   TextField "Text field_116" at 102,429 size 382x38; Text 'Tank 1P GTT Isolation Valve Feedback - Opened CV422'
   TextField "Text field_117" at 102,465 size 374x38; Text 'Tank 1P GTT Isolation Valve Feedback - Closed CV422'
   TextField "Text field_118" at 102,501 size 371x38; Text 'Tank 1P Tank Vent Valve 1 Feedback - Opened CV441-1PA'
   TextField "Text field_119" at 102,537 size 363x38; Text 'Tank 1P Tank Vent Valve 1 Feedback - Closed CV441-1PA'
   TextField "Text field_120" at 102,573 size 371x38; Text 'Tank 1P Tank Vent Valve 2 Feedback - Opened CV441-1PB'
   TextField "Text field_121" at 102,609 size 363x38; Text 'Tank 1P Tank Vent Valve 2 Feedback - Closed CV441-1PB'
   TextField "Text field_122" at 102,690 size 100x21; Text 'Spare Input'
   TextField "Text field_123" at 636,113 size 382x38; Text 'Tank 1S GTT Isolation Valve Feedback - Opened CV421'
   TextField "Text field_124" at 636,148 size 374x38; Text 'Tank 1S GTT Isolation Valve Feedback - Closed CV421'
   TextField "Text field_125" at 636,184 size 371x38; Text 'Tank 1S Tank Vent Valve 1 Feedback - Opened CV440-1SA'
   TextField "Text field_126" at 636,219 size 363x38; Text 'Tank 1S Tank Vent Valve 1 Feedback - Closed CV440-1SA'
   TextField "Text field_127" at 636,255 size 371x38; Text 'Tank 1S Tank Vent Valve 2 Feedback - Opened CV440-1SB'
   TextField "Text field_128" at 636,291 size 363x38; Text 'Tank 1S Tank Vent Valve 2 Feedback - Closed CV440-1SB'
   TextField "Text field_129" at 636,328 size 100x21; Text 'Spare Input'
   TextField "Text field_130" at 636,366 size 100x21; Text 'Spare Input'
   TextField "Text field_131" at 635,431 size 260x38; Text 'FPT BWT Level High High Switch LS425-FPT'
   TextField "Text field_132" at 635,467 size 270x38; Text 'RIO1 Tanks Pressure Switch Hi Hi PS436-FPT/1P/1S'
   TextField "Text field_133" at 635,503 size 294x38; Text 'Tank 1P BWT Level High High Switch LS425-1P'
   TextField "Text field_134" at 635,611 size 100x21; Text 'Spare Input'
   TextField "Text field_135" at 635,648 size 100x21; Text 'Spare Input'
   TextField "Text field_136" at 635,688 size 100x21; Text 'Spare Input'
   TextField "Text field_137" at 635,539 size 294x38; Text 'Tank 1S BWT Level High High Switch LS425-1S'
   TextField "Text field_138" at 635,576 size 100x21; Text 'Spare Input'
   TextField "Text field_115" at 102,654 size 100x21; Text 'Spare Input'
   AlarmView "Alarm view_1" at 0,777 size 1280x23
   Group "Group" at 455,41 size 373x50
   Button "HmiScreenItemData_8" at 469,45 size 355x40; TextOn 'Back'; TextOff 'Text'
      on Click: "TitleUpdater"()
   TextField "Screen title" at 455,41 size 373x50; Text 'Screen title'

screen "IGG Digital Outputs" 1280x800, template "Template"
   on GenerateScreen: "TitleUpdater"()
   Button "HmiScreenItemData_1" at 1,1 size 150x43; TextOn 'Back'; TextOff 'Commissioning'
      on Release: ActivateScreen("Commissioning Main Page", 0)
   AlarmView "Alarm view_1" at 0,777 size 1280x23
   TextField "Text field_1" at 395,239 size 55x22; Text 'Q0.0'
   TextField "Text field_2" at 395,290 size 55x22; Text 'Q0.1'
   TextField "Text field_3" at 395,342 size 55x22; Text 'Q0.2'
   TextField "Text field_4" at 395,394 size 55x22; Text 'Q0.3'
   TextField "Text field_5" at 395,446 size 55x22; Text 'Q0.4'
   TextField "Text field_6" at 395,498 size 55x22; Text 'Q0.5'
   TextField "Text field_7" at 395,550 size 55x22; Text 'Q0.6'
   TextField "Text field_8" at 395,602 size 55x22; Text 'Q0.7'
   Circle "Circle_1" at 455,239 size 20x20
      Appearance <- "14_DQ_Data_E500A_CNTRL"
   Circle "Circle_2" at 455,290 size 20x20
      Appearance <- "14_DQ_Data_E500B_CNTRL"
   Circle "Circle_3" at 455,342 size 20x20
      Appearance <- "14_DQ_Data_E139_CNTRL"
   Circle "Circle_4" at 455,394 size 20x20
      Appearance <- "14_DQ_Data_CV311_312_CNTRL"
   Circle "Circle_5" at 455,446 size 20x20
      Appearance <- "14_DQ_Data_CV321_322_CNTRL"
   Circle "Circle_6" at 455,498 size 20x20
      Appearance <- "14_DQ_Data_CV401_CNTRL"
   Circle "Circle_7" at 455,550 size 20x20
      Appearance <- "14_DQ_Data_CV431_432_CNTRL"
   Circle "Circle_8" at 455,602 size 20x20
      Appearance <- "14_DQ_Data_R2_SPR_DQ_0_7"
   TextField "Text field_9" at 412,206 size 49x26; Text 'Q0'
   TextField "Text field_10" at 698,239 size 55x22; Text 'Q1.0'
   TextField "Text field_11" at 698,290 size 55x22; Text 'Q1.1'
   TextField "Text field_12" at 698,342 size 55x22; Text 'Q1.2'
   TextField "Text field_13" at 698,394 size 55x22; Text 'Q1.3'
   TextField "Text field_14" at 698,446 size 55x22; Text 'Q1.4'
   TextField "Text field_15" at 698,498 size 55x22; Text 'Q1.5'
   TextField "Text field_16" at 698,550 size 55x22; Text 'Q1.6'
   TextField "Text field_17" at 698,602 size 55x22; Text 'Q1.7'
   Circle "Circle_9" at 758,239 size 20x20
      Appearance <- "14_DQ_Data_R2_SPR_DQ_1_0"
   Circle "Circle_10" at 758,290 size 20x20
      Appearance <- "14_DQ_Data_24K2"
   Circle "Circle_11" at 758,342 size 20x20
      Appearance <- "14_DQ_Data_24K3"
   Circle "Circle_12" at 758,394 size 20x20
      Appearance <- "14_DQ_Data_24K4"
   Circle "Circle_13" at 758,446 size 20x20
      Appearance <- "14_DQ_Data_24PF1"
   Circle "Circle_14" at 758,498 size 20x20
      Appearance <- "14_DQ_Data_24PF2"
   Circle "Circle_15" at 758,550 size 20x20
      Appearance <- "14_DQ_Data_24PF3"
   Circle "Circle_16" at 758,602 size 20x20
      Appearance <- "14_DQ_Data_24PF4"
   TextField "Text field_18" at 715,206 size 49x26; Text 'Q1'
   TextField "Text field_37" at 328,167 size 254x26; Text 'IGG System PLC (Rack 1)'
   Button "Button_9" at 330,493 size 60x35; TextOff 'Override'
      on Press: InvertBit("80_From_HMI_MAN_DQ_0_5")
      Visibility <- "82_To_HMI_CRNT_MODE_IGG"
   Button "Button_10" at 330,441 size 60x35; TextOff 'Override'
      on Press: InvertBit("80_From_HMI_MAN_DQ_0_4")
      Visibility <- "82_To_HMI_CRNT_MODE_IGG"
   Button "Button_11" at 330,388 size 60x35; TextOff 'Override'
      on Press: InvertBit("80_From_HMI_MAN_DQ_0_3")
      Visibility <- "82_To_HMI_CRNT_MODE_IGG"
   Button "Button_12" at 631,596 size 60x35; TextOff 'Override'
      on Press: InvertBit("80_From_HMI_MAN_DQ_1_7")
      Visibility <- "82_To_HMI_CRNT_MODE_IGG"
   Button "Button_14" at 631,283 size 60x35; TextOff 'Override'
      on Press: InvertBit("80_From_HMI_MAN_DQ_1_1")
      Visibility <- "82_To_HMI_CRNT_MODE_IGG"
   TextField "Text field_56" at 481,239 size 140x22; Text 'Fuel Pump 1 E500A'
   TextField "Text field_57" at 481,290 size 140x22; Text 'Fuel Pump 2 E500B'
   TextField "Text field_58" at 481,342 size 140x22; Text 'CA Blower E139'
   TextField "Text field_59" at 481,394 size 140x22; Text 'CSW Inlet Valves CV311'
   TextField "Text field_60" at 481,446 size 140x22; Text 'CSW Drain Valves CV322'
   TextField "Text field_61" at 481,498 size 140x22; Text 'IG Supply Valve CV401'
   TextField "Text field_62" at 481,549 size 140x22; Text 'CB/BWTS Valve CV432'
   TextField "Text field_63" at 481,602 size 140x22; Text 'Spare Output'
   TextField "Text field_64" at 786,242 size 140x22; Text 'Spare Output'
   TextField "Text field_65" at 786,290 size 140x22; Text 'Atmospheric Alarm'
   TextField "Text field_66" at 786,342 size 140x22; Text 'IGG Shutdown Alarm'
   TextField "Text field_67" at 786,394 size 140x22; Text 'IGG Warning Alarm'
   TextField "Text field_68" at 786,446 size 140x22; Text 'IGG Running'
   TextField "Text field_69" at 786,497 size 140x22; Text 'Shutdown Alarm'
   TextField "Text field_70" at 786,550 size 140x22; Text 'Warning Alarm'
   TextField "Text field_71" at 786,602 size 140x22; Text 'Buzzer'
   Button "Button_15" at 330,336 size 60x35; TextOff 'Override'
      on Press: InvertBit("80_From_HMI_MAN_DQ_0_2")
      Visibility <- "82_To_HMI_CRNT_MODE_IGG"
   Button "Button_16" at 330,283 size 60x35; TextOff 'Override'
      on Press: InvertBit("80_From_HMI_MAN_DQ_0_1")
      Visibility <- "82_To_HMI_CRNT_MODE_IGG"
   Button "Button_17" at 330,546 size 60x35; TextOff 'Override'
      on Press: InvertBit("80_From_HMI_MAN_DQ_0_6")
      Visibility <- "82_To_HMI_CRNT_MODE_IGG"
   Button "Button_18" at 330,599 size 60x35; TextOff 'Override'
      on Press: InvertBit("80_From_HMI_MAN_DQ_0_7(1)")
      Visibility <- "82_To_HMI_CRNT_MODE_IGG"
   Button "Button_19" at 330,231 size 60x35; TextOff 'Override'
      on Press: InvertBit("80_From_HMI_MAN_DQ_0_0")
      Visibility <- "82_To_HMI_CRNT_MODE_IGG"
   Button "Button_20" at 631,231 size 60x35; TextOff 'Override'
      on Press: InvertBit("80_From_HMI_MAN_DQ_1_0(1)")
      Visibility <- "82_To_HMI_CRNT_MODE_IGG"
   Button "Button_21" at 631,335 size 60x35; TextOff 'Override'
      on Press: InvertBit("80_From_HMI_MAN_DQ_1_2")
      Visibility <- "82_To_HMI_CRNT_MODE_IGG"
   Button "Button_22" at 631,387 size 60x35; TextOff 'Override'
      on Press: InvertBit("80_From_HMI_MAN_DQ_1_3")
      Visibility <- "82_To_HMI_CRNT_MODE_IGG"
   Button "Button_23" at 631,439 size 60x35; TextOff 'Override'
      on Press: InvertBit("80_From_HMI_MAN_DQ_1_4")
      Visibility <- "82_To_HMI_CRNT_MODE_IGG"
   Button "Button_24" at 631,491 size 60x35; TextOff 'Override'
      on Press: InvertBit("80_From_HMI_MAN_DQ_1_5")
      Visibility <- "82_To_HMI_CRNT_MODE_IGG"
   Button "Button_25" at 631,543 size 60x35; TextOff 'Override'
      on Press: InvertBit("80_From_HMI_MAN_DQ_1_6(1)")
      Visibility <- "82_To_HMI_CRNT_MODE_IGG"
   Group "Group" at 455,41 size 373x50
   Button "HmiScreenItemData_8" at 469,45 size 355x40; TextOn 'Back'; TextOff 'Text'
   TextField "Screen title" at 455,41 size 373x50; Text 'Screen title'

screen "BWT Digital Outputs" 1280x800, template "Template"
   on GenerateScreen: "TitleUpdater"()
   TextField "Text field_1" at 79,178 size 55x22; Text 'Q0.0'
   TextField "Text field_2" at 79,229 size 55x22; Text 'Q0.1'
   TextField "Text field_3" at 79,281 size 55x22; Text 'Q0.2'
   TextField "Text field_4" at 79,333 size 55x22; Text 'Q0.3'
   TextField "Text field_5" at 79,385 size 55x22; Text 'Q0.4'
   TextField "Text field_6" at 79,437 size 55x22; Text 'Q0.5'
   TextField "Text field_7" at 79,489 size 55x22; Text 'Q0.6'
   TextField "Text field_8" at 79,541 size 55x22; Text 'Q0.7'
   Circle "Circle_1" at 139,178 size 20x20
      Appearance <- "14_DQ_Data_E500A_CNTRL"
   Circle "Circle_2" at 139,229 size 20x20
      Appearance <- "14_DQ_Data_E500B_CNTRL"
   Circle "Circle_3" at 139,281 size 20x20
      Appearance <- "14_DQ_Data_E139_CNTRL"
   Circle "Circle_4" at 139,333 size 20x20
      Appearance <- "14_DQ_Data_CV311_312_CNTRL"
   Circle "Circle_5" at 139,385 size 20x20
      Appearance <- "14_DQ_Data_CV321_322_CNTRL"
   Circle "Circle_6" at 139,437 size 20x20
      Appearance <- "14_DQ_Data_CV401_CNTRL"
   Circle "Circle_7" at 139,489 size 20x20
      Appearance <- "14_DQ_Data_CV431_432_CNTRL"
   Circle "Circle_8" at 139,541 size 20x20
      Appearance <- "14_DQ_Data_R2_SPR_DQ_0_7"
   TextField "Text field_9" at 96,145 size 49x26; Text 'Q0'
   TextField "Text field_10" at 382,178 size 55x22; Text 'Q1.0'
   TextField "Text field_11" at 382,229 size 55x22; Text 'Q1.1'
   TextField "Text field_12" at 382,281 size 55x22; Text 'Q1.2'
   TextField "Text field_13" at 382,333 size 55x22; Text 'Q1.3'
   TextField "Text field_14" at 382,385 size 55x22; Text 'Q1.4'
   TextField "Text field_15" at 382,437 size 55x22; Text 'Q1.5'
   TextField "Text field_16" at 382,489 size 55x22; Text 'Q1.6'
   TextField "Text field_17" at 382,541 size 55x22; Text 'Q1.7'
   Circle "Circle_9" at 442,178 size 20x20
      Appearance <- "14_DQ_Data_R2_SPR_DQ_1_0"
   Circle "Circle_10" at 442,229 size 20x20
      Appearance <- "14_DQ_Data_24K2"
   Circle "Circle_11" at 442,281 size 20x20
      Appearance <- "14_DQ_Data_24K3"
   Circle "Circle_12" at 442,333 size 20x20
      Appearance <- "14_DQ_Data_24K4"
   Circle "Circle_13" at 442,385 size 20x20
      Appearance <- "14_DQ_Data_24PF1"
   Circle "Circle_14" at 442,437 size 20x20
      Appearance <- "14_DQ_Data_24PF2"
   Circle "Circle_15" at 442,489 size 20x20
      Appearance <- "14_DQ_Data_24PF3"
   Circle "Circle_16" at 442,541 size 20x20
      Appearance <- "14_DQ_Data_24PF4"
   TextField "Text field_18" at 399,145 size 49x26; Text 'Q1'
   TextField "Text field_37" at 12,106 size 263x26; Text 'BWT Control PLC (Rack 3)'
   Button "HmiScreenItemData_1" at 1,1 size 150x43; TextOn 'Back'; TextOff 'Commissioning'
      on Release: ActivateScreen("Commissioning Main Page", 0)
   Button "Button_9" at 14,432 size 60x35; TextOff 'Override'
      on Press: InvertBit("80_From_HMI_MAN_DQ_0_5")
      Visibility <- "82_To_HMI_CRNT_MODE_IGG"
   Button "Button_10" at 14,380 size 60x35; TextOff 'Override'
      on Press: InvertBit("80_From_HMI_MAN_DQ_0_4")
      Visibility <- "82_To_HMI_CRNT_MODE_IGG"
   Button "Button_11" at 14,327 size 60x35; TextOff 'Override'
      on Press: InvertBit("80_From_HMI_MAN_DQ_0_3")
      Visibility <- "82_To_HMI_CRNT_MODE_IGG"
   Button "Button_12" at 315,535 size 60x35; TextOff 'Override'
      on Press: InvertBit("80_From_HMI_MAN_DQ_1_7")
      Visibility <- "82_To_HMI_CRNT_MODE_IGG"
   Button "Button_14" at 315,222 size 60x35; TextOff 'Override'
      on Press: InvertBit("80_From_HMI_MAN_DQ_1_1")
      Visibility <- "82_To_HMI_CRNT_MODE_IGG"
   TextField "Text field_56" at 165,174 size 117x42; Text 'Fuel Pump 1 E500A'
   TextField "Text field_57" at 165,223 size 117x42; Text 'Fuel Pump 2 E500B'
   TextField "Text field_58" at 165,277 size 100x42; Text 'CA Blower E139'
   TextField "Text field_59" at 165,327 size 161x42; Text 'CSW Inlet Valves CV311'
   TextField "Text field_60" at 165,378 size 166x42; Text 'CSW Drain Valves CV322'
   TextField "Text field_61" at 165,434 size 149x42; Text 'IG Supply Valve CV401'
   TextField "Text field_62" at 165,489 size 154x42; Text 'CB/BWTS Valve CV432'
   TextField "Text field_63" at 165,538 size 125x23; Text 'Spare Output'
   TextField "Text field_64" at 470,175 size 125x23; Text 'Spare Output'
   TextField "Text field_65" at 470,224 size 178x23; Text 'Atmospheric Alarm'
   TextField "Text field_66" at 470,278 size 194x23; Text 'IGG Shutdown Alarm'
   TextField "Text field_67" at 470,328 size 180x23; Text 'IGG Warning Alarm'
   TextField "Text field_68" at 470,379 size 119x23; Text 'IGG Running'
   TextField "Text field_69" at 470,431 size 154x23; Text 'Shutdown Alarm'
   TextField "Text field_70" at 470,490 size 140x23; Text 'Warning Alarm'
   TextField "Text field_71" at 470,539 size 67x23; Text 'Buzzer'
   Button "Button_15" at 14,275 size 60x35; TextOff 'Override'
      on Press: InvertBit("80_From_HMI_MAN_DQ_0_2")
      Visibility <- "82_To_HMI_CRNT_MODE_IGG"
   Button "Button_16" at 14,222 size 60x35; TextOff 'Override'
      on Press: InvertBit("80_From_HMI_MAN_DQ_0_1")
      Visibility <- "82_To_HMI_CRNT_MODE_IGG"
   Button "Button_17" at 14,485 size 60x35; TextOff 'Override'
      on Press: InvertBit("80_From_HMI_MAN_DQ_0_6")
      Visibility <- "82_To_HMI_CRNT_MODE_IGG"
   Button "Button_18" at 14,538 size 60x35; TextOff 'Override'
      on Press: InvertBit("80_From_HMI_MAN_DQ_0_7(1)")
      Visibility <- "82_To_HMI_CRNT_MODE_IGG"
   Button "Button_19" at 14,170 size 60x35; TextOff 'Override'
      on Press: InvertBit("80_From_HMI_MAN_DQ_0_0")
      Visibility <- "82_To_HMI_CRNT_MODE_IGG"
   Button "Button_20" at 315,170 size 60x35; TextOff 'Override'
      on Press: InvertBit("80_From_HMI_MAN_DQ_1_0(1)")
      Visibility <- "82_To_HMI_CRNT_MODE_IGG"
   Button "Button_21" at 315,274 size 60x35; TextOff 'Override'
      on Press: InvertBit("80_From_HMI_MAN_DQ_1_2")
      Visibility <- "82_To_HMI_CRNT_MODE_IGG"
   Button "Button_22" at 315,326 size 60x35; TextOff 'Override'
      on Press: InvertBit("80_From_HMI_MAN_DQ_1_3")
      Visibility <- "82_To_HMI_CRNT_MODE_IGG"
   Button "Button_23" at 315,378 size 60x35; TextOff 'Override'
      on Press: InvertBit("80_From_HMI_MAN_DQ_1_4")
      Visibility <- "82_To_HMI_CRNT_MODE_IGG"
   Button "Button_24" at 315,430 size 60x35; TextOff 'Override'
      on Press: InvertBit("80_From_HMI_MAN_DQ_1_5")
      Visibility <- "82_To_HMI_CRNT_MODE_IGG"
   Button "Button_25" at 315,482 size 60x35; TextOff 'Override'
      on Press: InvertBit("80_From_HMI_MAN_DQ_1_6(1)")
      Visibility <- "82_To_HMI_CRNT_MODE_IGG"
   AlarmView "Alarm view_1" at 0,777 size 1280x23
   TextField "Text field_19" at 23,309 size 1188x123; Text 'Re - Work Required Througout This page'
   Group "Group" at 455,41 size 373x50
   Button "HmiScreenItemData_8" at 469,45 size 355x40; TextOn 'Back'; TextOff 'Text'
   TextField "Screen title" at 455,41 size 373x50; Text 'Screen title'

screen "BWT Analogue Inputs" 1280x800, template "Template"
   on GenerateScreen: "TitleUpdater"()
   IOField "I/O field_62" at 1208,191 size 60x22; FormatPattern 99.9
   IOField "I/O field_61" at 1140,191 size 60x22; FormatPattern 99.9
   Button "HmiScreenItemData_1" at 1,1 size 150x43; TextOn 'Back'; TextOff 'Commissioning'
      on Release: ActivateScreen("Commissioning Main Page", 0)
   TextField "Text field_82" at 60,150 size 220x22; Text 'PIT-102 - CA Pressure (Pre-Ignition)'
   TextField "Text field_90" at 286,124 size 64x20; Text 'Reading'
   IOField "I/O field_2" at 287,150 size 70x22; FormatPattern 9999; Unit  mBar
      ProcessValue <- "12_AI_Data_PIT102_SCALED(1)"
   TextField "Text field_1" at 359,124 size 68x20; Text 'Low Low'
   IOField "I/O field_1" at 361,150 size 60x22; Authorization "Parameter Change"; FormatPattern 9999
      ProcessValue <- "84_Setpoints_PIT102_Pilot_LowLow"
   TextField "Text field_2" at 442,124 size 37x20; Text 'Low'
   IOField "I/O field_3" at 429,150 size 60x22; Authorization "Parameter Change"; FormatPattern 9999
      ProcessValue <- "84_Setpoints_PIT102_Pilot_Low"
   TextField "Text field_3" at 509,124 size 37x20; Text 'High'
   IOField "I/O field_4" at 497,150 size 60x22; Authorization "Parameter Change"; FormatPattern 9999
      ProcessValue <- "84_Setpoints_PIT102_Pilot_High"
   TextField "Text field_4" at 561,124 size 74x20; Text 'High High'
   IOField "I/O field_5" at 565,150 size 60x22; Authorization "Parameter Change"; FormatPattern 9999
      ProcessValue <- "84_Setpoints_PIT102_Pilot_HighHigh"
   TextField "Text field_5" at 434,100 size 76x20; Text 'Setpoints'
   TextField "Text field_6" at 7,150 size 53x22; Text 'IW112'
   TextField "Text field_7" at 60,270 size 220x22; Text 'TIT-401 - IG Temperature'
   IOField "I/O field_6" at 287,270 size 70x22; FormatPattern s999.9; Unit  °C
      ProcessValue <- "12_AI_Data_TIT401_SCALED"
   IOField "I/O field_7" at 361,270 size 60x22; FormatPattern s999.9
   IOField "I/O field_8" at 429,270 size 60x22; FormatPattern s999.9
   IOField "I/O field_9" at 497,270 size 60x22; Authorization "Parameter Change"; FormatPattern s999.9
      ProcessValue <- "84_Setpoints_TIT401_High"
   IOField "I/O field_10" at 565,270 size 60x22; Authorization "Parameter Change"; FormatPattern s999.9
      ProcessValue <- "84_Setpoints_TIT401_HighHigh"
   TextField "Text field_8" at 7,270 size 53x22; Text 'IW114'
   TextField "Text field_9" at 60,310 size 220x22; Text 'PIT-402 - IG Outlet Pres. (Pre-Ignitn.)'
   IOField "I/O field_11" at 287,310 size 70x22; FormatPattern 9999; Unit  mBar
      ProcessValue <- "12_AI_Data_PIT402_SCALED"
   IOField "I/O field_12" at 361,310 size 60x22; Authorization "Parameter Change"; FormatPattern 9999
      ProcessValue <- "84_Setpoints_PIT402_Pilot_LowLow"
   IOField "I/O field_13" at 429,310 size 60x22; Authorization "Parameter Change"; FormatPattern 9999
      ProcessValue <- "84_Setpoints_PIT402_Pilot_Low"
   IOField "I/O field_14" at 497,310 size 60x22; Authorization "Parameter Change"; FormatPattern 9999
      ProcessValue <- "84_Setpoints_PIT402_Pilot_High"
   IOField "I/O field_15" at 565,310 size 60x22; Authorization "Parameter Change"; FormatPattern 9999
      ProcessValue <- "84_Setpoints_PIT402_Pilot_HighHigh"
   TextField "Text field_10" at 7,310 size 53x22; Text 'IW116'
   TextField "Text field_11" at 60,430 size 220x22; Text 'CV-403 - IG Vent Valve Position Fbk'
   IOField "I/O field_16" at 287,430 size 70x22; FormatPattern 999; Unit  %
      ProcessValue <- "12_AI_Data_CV403_SCALED"
   IOField "I/O field_17" at 361,430 size 60x22; FormatPattern 999
   IOField "I/O field_18" at 429,430 size 60x22; FormatPattern 999
   IOField "I/O field_19" at 497,430 size 60x22; FormatPattern 999
   IOField "I/O field_20" at 565,430 size 60x22; FormatPattern 999
   TextField "Text field_12" at 7,430 size 53x22; Text 'IW118'
   TextField "Text field_13" at 60,470 size 220x22; Text 'CA Blower RPM'
   IOField "I/O field_21" at 287,470 size 70x22; FormatPattern 9999; Unit  RPM
      ProcessValue <- "12_AI_Data_E139_RPM_SCALED"
   IOField "I/O field_22" at 361,470 size 60x22; FormatPattern 9999
   IOField "I/O field_23" at 429,470 size 60x22; FormatPattern 9999
   IOField "I/O field_24" at 497,470 size 60x22; FormatPattern 9999
   IOField "I/O field_25" at 565,470 size 60x22; FormatPattern 9999
   TextField "Text field_14" at 7,470 size 54x22; Text 'IW120'
   TextField "Text field_15" at 61,511 size 220x22; Text 'CA Blower Current'
   IOField "I/O field_26" at 288,511 size 70x22; FormatPattern 999.9; Unit  A
      ProcessValue <- "12_AI_Data_E139_AMPS_SCALED"
   IOField "I/O field_27" at 362,511 size 60x22; FormatPattern 9999
   IOField "I/O field_28" at 430,511 size 60x22; FormatPattern 9999
   TextField "Text field_16" at 8,511 size 54x22; Text 'IW122'
   TextField "Text field_17" at 61,552 size 220x22; Text 'LIT-305 - FW Bulk Tank Level'
   IOField "I/O field_31" at 288,552 size 70x22; FormatPattern 99.9; Unit  %
      ProcessValue <- "12_AI_Data_LIT305_SCALED"
   TextField "Text field_18" at 8,552 size 53x22; Text 'IW124'
   TextField "Text field_19" at 61,592 size 220x22; Text 'Spare'
   IOField "I/O field_36" at 288,592 size 70x22; FormatPattern 9.9; Unit  
      ProcessValue <- "12_AI_Data_R1_SPR_AI_126_SCALED"
   IOField "I/O field_37" at 362,592 size 60x22; FormatPattern 9.9
   IOField "I/O field_38" at 430,592 size 60x22; FormatPattern 9.9
   IOField "I/O field_39" at 498,592 size 60x22; FormatPattern 9.9
   IOField "I/O field_40" at 566,592 size 60x22; FormatPattern 9.9
   TextField "Text field_20" at 8,592 size 53x22; Text 'IW126'
   TextField "Text field_21" at 703,151 size 220x22; Text 'Atmospheric Oxygen 1'
   IOField "I/O field_41" at 930,151 size 70x22; FormatPattern 99.99; Unit %
      ProcessValue <- "12_AI_Data_AT_O2_01_SCALED"
   IOField "I/O field_42" at 1004,151 size 60x22; Authorization "Commissioning"; FormatPattern 99.9
      ProcessValue <- "84_Setpoints_AT_O2_1_LowLow"
   IOField "I/O field_43" at 1072,151 size 60x22; Authorization "Commissioning"; FormatPattern 99.9
      ProcessValue <- "84_Setpoints_AT_O2_1_Low"
   IOField "I/O field_44" at 1140,151 size 60x22; FormatPattern 99.9
   IOField "I/O field_45" at 1208,151 size 60x22; FormatPattern 99.9
   TextField "Text field_22" at 650,151 size 53x22; Text 'IW128'
   TextField "Text field_23" at 703,191 size 220x22; Text 'Atmospheric Oxygen 2'
   IOField "I/O field_46" at 930,191 size 70x22; FormatPattern 99.99; Unit %
      ProcessValue <- "12_AI_Data_AT_O2_02_SCALED"
   TextField "Text field_24" at 650,191 size 53x22; Text 'IW130'
   TextField "Text field_26" at 928,124 size 64x20; Text 'Reading'
   TextField "Text field_27" at 1001,124 size 68x20; Text 'Low Low'
   TextField "Text field_28" at 1082,124 size 37x20; Text 'Low'
   TextField "Text field_29" at 1150,124 size 37x20; Text 'High'
   TextField "Text field_30" at 1203,124 size 74x20; Text 'High High'
   TextField "Text field_31" at 1076,100 size 76x20; Text 'Setpoints'
   TextField "Text field_51" at 703,231 size 220x22; Text 'Spare'
   IOField "I/O field_101" at 930,231 size 70x22; FormatPattern 99.9
      ProcessValue <- "12_AI_Data_R1_SPR_AI_132_SCALED"
   TextField "Text field_56" at 650,231 size 53x22; Text 'IW132'
   TextField "Text field_57" at 703,271 size 220x22; Text 'TIT-315 - Shell CSW Temperature'
   IOField "I/O field_106" at 930,271 size 70x22; FormatPattern s999.9; Unit  °C
      ProcessValue <- "12_AI_Data_TIT315_SCALED"
   IOField "I/O field_107" at 1004,271 size 60x22; FormatPattern s999.9
   IOField "I/O field_108" at 1072,271 size 60x22; FormatPattern s999.9
   TextField "Text field_58" at 650,271 size 54x22; Text 'IW134'
   TextField "Text field_59" at 703,311 size 220x22; Text 'TIT-319 - Inlet CSW Temperature'
   IOField "I/O field_111" at 930,311 size 70x22; FormatPattern s999.9; Unit  °C
      ProcessValue <- "12_AI_Data_TIT319_SCALED"
   IOField "I/O field_112" at 1004,311 size 60x22; FormatPattern s999.9
   IOField "I/O field_113" at 1072,311 size 60x22; FormatPattern s999.9
   TextField "Text field_60" at 650,311 size 53x22; Text 'IW136'
   TextField "Text field_61" at 703,351 size 220x22; Text 'TIT-360 - Outlet CSW Temperature'
   IOField "I/O field_116" at 930,351 size 70x22; FormatPattern s999.9; Unit  °C
      ProcessValue <- "12_AI_Data_TIT360_SCALED"
   IOField "I/O field_117" at 1004,351 size 60x22; FormatPattern s999.9
   IOField "I/O field_118" at 1072,351 size 60x22; FormatPattern s999.9
   TextField "Text field_62" at 650,351 size 53x22; Text 'IW138'
   TextField "Text field_63" at 703,391 size 220x22; Text 'PIT-359 - Inlet CSW Pressure'
   IOField "I/O field_121" at 930,391 size 70x22; FormatPattern 99.9; Unit  Bar
      ProcessValue <- "12_AI_Data_PIT359_SCALED"
   TextField "Text field_64" at 650,391 size 53x22; Text 'IW140'
   TextField "Text field_41" at 133,124 size 89x20; Text 'Description'
   TextField "Text field_42" at 771,124 size 89x20; Text 'Description'
   TextField "Text field_43" at 17,124 size 37x20; Text 'AI'
   TextField "Text field_44" at 661,124 size 37x20; Text 'AI'
   TextField "Text field_47" at 702,431 size 220x22; Text 'PIT-316 - Outlet CSW Pressure'
   IOField "I/O field_81" at 929,431 size 70x22; FormatPattern 99.9; Unit  Bar
      ProcessValue <- "12_AI_Data_PIT316_SCALED"
   TextField "Text field_48" at 649,431 size 53x22; Text 'IW142'
   IOField "I/O field_109" at 1140,271 size 60x22; Authorization "Parameter Change"; FormatPattern s999.9
      ProcessValue <- "84_Setpoints_TIT315_High"
   IOField "I/O field_110" at 1208,271 size 60x22; Authorization "Parameter Change"; FormatPattern s999.9
      ProcessValue <- "84_Setpoints_TIT315_HighHigh"
   IOField "I/O field_114" at 1140,311 size 60x22; Authorization "Parameter Change"; FormatPattern s999.9
      ProcessValue <- "84_Setpoints_TIT319_High"
   IOField "I/O field_115" at 1208,311 size 60x22; Authorization "Parameter Change"; FormatPattern s999.9
      ProcessValue <- "84_Setpoints_TIT319_HighHigh"
   IOField "I/O field_119" at 1140,351 size 60x22; Authorization "Parameter Change"; FormatPattern s999.9
      ProcessValue <- "84_Setpoints_TIT360_High"
   IOField "I/O field_120" at 1208,351 size 60x22; Authorization "Parameter Change"; FormatPattern s999.9
      ProcessValue <- "84_Setpoints_TIT360_HighHigh"
   IOField "I/O field_124" at 1140,391 size 60x22; Authorization "Parameter Change"; FormatPattern 99.9
      ProcessValue <- "84_Setpoints_PIT359_High"
   IOField "I/O field_125" at 1208,391 size 60x22; Authorization "Parameter Change"; FormatPattern 99.9
      ProcessValue <- "84_Setpoints_PIT359_HighHigh"
   IOField "I/O field_84" at 1139,431 size 60x22; Authorization "Parameter Change"; FormatPattern 99.9
      ProcessValue <- "84_Setpoints_PIT316_High"
   IOField "I/O field_85" at 1207,431 size 60x22; Authorization "Parameter Change"; FormatPattern 99.9
      ProcessValue <- "84_Setpoints_PIT316_HighHigh"
   IOField "I/O field_122" at 1004,391 size 60x22; Authorization "Parameter Change"; FormatPattern 99.9
      ProcessValue <- "84_Setpoints_PIT359_LowLow"
   IOField "I/O field_123" at 1072,391 size 60x22; Authorization "Parameter Change"; FormatPattern 99.9
      ProcessValue <- "84_Setpoints_PIT359_Low"
   IOField "I/O field_82" at 1003,431 size 60x22; Authorization "Parameter Change"; FormatPattern 99.9
      ProcessValue <- "84_Setpoints_PIT316_LowLow"
   IOField "I/O field_83" at 1071,431 size 60x22; Authorization "Parameter Change"; FormatPattern 99.9
      ProcessValue <- "84_Setpoints_PIT316_Low"
   TextField "Text field_52" at 17,91 size 340x26; Text 'BWT Control System PLC (Rack 3)'
   TextField "Text field_54" at 649,719 size 228x62; Text 'Note: CSW = Cooling Sea Water'
   Button "Button_1" at 1160,732 size 100x35; TextOn 'BWTS Digital Inputs.'; TextOff 'Next'
      on Click: ActivateScreen("BC Analogue Inputs", 0)
   TextField "Text field_25" at 60,231 size 220x22; Text 'PIT-102 - CA Pressure (Post-Ignition)'
   IOField "I/O field_52" at 361,231 size 60x22; Authorization "Parameter Change"; FormatPattern 9999
      ProcessValue <- "84_Setpoints_PIT102_Post_LowLow"
   IOField "I/O field_53" at 429,231 size 60x22; Authorization "Parameter Change"; FormatPattern 9999
      ProcessValue <- "84_Setpoints_PIT102_Post_Low"
   IOField "I/O field_54" at 497,231 size 60x22; Authorization "Parameter Change"; FormatPattern 9999
      ProcessValue <- "84_Setpoints_PIT102_Post_High"
   IOField "I/O field_55" at 565,231 size 60x22; Authorization "Parameter Change"; FormatPattern 9999
      ProcessValue <- "84_Setpoints_PIT102_Post_HighHigh"
   TextField "Text field_32" at 7,231 size 53x22; Text 'IW112'
   TextField "Text field_33" at 60,391 size 220x22; Text 'PIT-402 - IG Outlet Pres. (Post-Ignitn)'
   IOField "I/O field_57" at 361,391 size 60x22; Authorization "Parameter Change"; FormatPattern 9999
      ProcessValue <- "84_Setpoints_PIT402_Post_LowLow"
   IOField "I/O field_58" at 429,391 size 60x22; Authorization "Parameter Change"; FormatPattern 9999
      ProcessValue <- "84_Setpoints_PIT402_Post_Low"
   IOField "I/O field_59" at 497,391 size 60x22; Authorization "Parameter Change"; FormatPattern 9999
      ProcessValue <- "84_Setpoints_PIT402_Post_High"
   IOField "I/O field_60" at 565,391 size 60x22; Authorization "Parameter Change"; FormatPattern 9999
      ProcessValue <- "84_Setpoints_PIT402_Post_HighHigh"
   TextField "Text field_34" at 7,391 size 53x22; Text 'IW116'
   IOField "I/O field_47" at 1004,191 size 60x22; Authorization "Commissioning"; FormatPattern 99.9
      ProcessValue <- "84_Setpoints_AT_O2_2_LowLow"
   IOField "I/O field_48" at 1072,191 size 60x22; Authorization "Commissioning"; FormatPattern 99.9
      ProcessValue <- "84_Setpoints_AT_O2_2_Low"
   TextField "Text field_35" at 61,191 size 220x22; Text 'PIT-102 - CA Pressure (Main)'
   IOField "I/O field_50" at 362,191 size 60x22; Authorization "Parameter Change"; FormatPattern 9999
      ProcessValue <- "84_Setpoints_PIT102_Main_LowLow"
   IOField "I/O field_63" at 430,191 size 60x22; Authorization "Parameter Change"; FormatPattern 9999
      ProcessValue <- "84_Setpoints_PIT102_Main_Low"
   IOField "I/O field_64" at 498,191 size 60x22; Authorization "Parameter Change"; FormatPattern 9999
      ProcessValue <- "84_Setpoints_PIT102_Main_High"
   IOField "I/O field_65" at 566,191 size 60x22; Authorization "Parameter Change"; FormatPattern 9999
      ProcessValue <- "84_Setpoints_PIT102_Main_HighHigh"
   TextField "Text field_36" at 8,191 size 53x22; Text 'IW112'
   IOField "I/O field_49" at 1004,231 size 60x22; FormatPattern 999
   IOField "I/O field_51" at 1072,231 size 60x22; FormatPattern 999
   IOField "I/O field_66" at 1140,231 size 60x22; FormatPattern 999
   IOField "I/O field_67" at 1208,231 size 60x22; FormatPattern 999
   TextField "Text field_37" at 61,349 size 220x22; Text 'PIT-402 - IG Outlet Pres. (Main)'
   IOField "I/O field_69" at 362,349 size 60x22; Authorization "Parameter Change"; FormatPattern 9999
      ProcessValue <- "84_Setpoints_PIT402_Main_LowLow"
   IOField "I/O field_70" at 430,349 size 60x22; Authorization "Parameter Change"; FormatPattern 9999
      ProcessValue <- "84_Setpoints_PIT402_Main_Low"
   IOField "I/O field_71" at 498,349 size 60x22; Authorization "Parameter Change"; FormatPattern 9999
      ProcessValue <- "84_Setpoints_PIT402_Main_High"
   IOField "I/O field_72" at 566,349 size 60x22; Authorization "Parameter Change"; FormatPattern 9999
      ProcessValue <- "84_Setpoints_PIT402_Main_HighHigh"
   TextField "Text field_38" at 8,349 size 53x22; Text 'IW116'
   IOField "I/O field_29" at 566,511 size 60x22; FormatPattern 9999
   IOField "I/O field_30" at 499,511 size 60x22; FormatPattern 9999
   IOField "I/O field_32" at 361,552 size 60x22; FormatPattern 9999
   IOField "I/O field_33" at 429,552 size 60x22; FormatPattern 9999
   IOField "I/O field_34" at 565,552 size 60x22; FormatPattern 9999
   IOField "I/O field_35" at 498,552 size 60x22; FormatPattern 9999
   TextField "Text field_39" at 1109,687 size 151x62; Text 'To BC Analogue Inputs'
   AlarmView "Alarm view_1" at 0,777 size 1280x23
   TextField "Text field_40" at 23,309 size 1188x123; Text 'Re - Work Required Througout This page'
   Group "Group" at 455,41 size 373x50
   Button "HmiScreenItemData_8" at 469,45 size 355x40; TextOn 'Back'; TextOff 'Text'
   TextField "Screen title" at 455,41 size 373x50; Text 'Screen title'

screen "BC Analogue Outputs" 1280x800, template "Template"
   on GenerateScreen: "TitleUpdater"()
   Button "HmiScreenItemData_1" at 1,1 size 150x43; TextOn 'Back'; TextOff 'Commissioning'
      on Release: ActivateScreen("Commissioning Main Page", 0)
   Button "Button_15" at 34,732 size 100x35; TextOn 'BWTS Digital Inputs'; TextOff 'Back'
      on Click: ActivateScreen("BC Analogue Inputs", 0)
   AlarmView "Alarm view_1" at 0,777 size 1280x23
   TextField "Text field_90" at 750,328 size 64x20; Text 'Reading'
   TextField "Text field_41" at 553,328 size 89x20; Text 'Description'
   TextField "Text field_43" at 437,328 size 37x20; Text 'AO'
   TextField "Text field_52" at 437,295 size 364x26; Text 'Burner Control System PLC (Rack 2)'
   TextField "Text field_4" at 481,444 size 220x22; Text 'Main Fuel Reg Valve Control'
   IOField "I/O field_4" at 749,446 size 70x22; FormatPattern 9999; Unit %
      ProcessValue <- "16_AQ_Data_CV203_CNTRL"
   TextField "Text field_8" at 428,444 size 53x22; Text 'QW100'
   TextField "Text field_9" at 481,368 size 220x22; Text 'Spare'
   TextField "Text field_12" at 480,482 size 220x22; Text 'Main Atom Air Reg Valve Control'
   IOField "I/O field_5" at 749,481 size 70x22; FormatPattern 9999; Unit %
      ProcessValue <- "16_AQ_Data_CV111_CNTRL"
   TextField "Text field_13" at 427,482 size 53x22; Text 'QW102'
   Button "Button_7" at 716,442 size 29x26; TextOff '+'
      on Press: function_b14e0dd5("80_From_HMI_MAN_AQ_INC_100(1)", 0)
      Visibility <- "82_To_HMI_CRNT_MODE_IGG"
   Button "Button_8" at 824,442 size 29x26; TextOff '-'
      on Press: function_b14e0dd5("80_From_HMI_MAN_AQ_DEC_100(1)", 0)
      Visibility <- "82_To_HMI_CRNT_MODE_IGG"
   Button "Button_9" at 716,480 size 29x26; TextOff '+'
      on Press: function_b14e0dd5("80_From_HMI_MAN_AQ_INC_102", 0)
      Visibility <- "82_To_HMI_CRNT_MODE_IGG"
   Button "Button_10" at 824,480 size 29x26; TextOff '-'
      on Press: function_b14e0dd5("80_From_HMI_MAN_AQ_DEC_102", 0)
      Visibility <- "82_To_HMI_CRNT_MODE_IGG"
   Button "Button_11" at 716,364 size 29x26; TextOff '+'
      on Click: SetBit("80_From_HMI_MAN_AQ_INC_96")
      Visibility <- "82_To_HMI_CRNT_MODE_IGG"
   Button "Button_12" at 824,364 size 29x26; TextOff '-'
      on Click: SetBit("80_From_HMI_MAN_AQ_DEC_96")
      Visibility <- "82_To_HMI_CRNT_MODE_IGG"
   Button "Button_13" at 716,405 size 29x26; TextOff '+'
      on Click: SetBit("80_From_HMI_MAN_AQ_INC_98")
      Visibility <- "82_To_HMI_CRNT_MODE_IGG"
   Button "Button_14" at 824,405 size 29x26; TextOff '-'
      on Click: SetBit("80_From_HMI_MAN_AQ_DEC_98")
      Visibility <- "82_To_HMI_CRNT_MODE_IGG"
   IOField "I/O field_6" at 749,368 size 70x22; FormatPattern 9.9; Unit  
      ProcessValue <- "16_AQ_Data_R2_SPR_AQ_96"
   IOField "I/O field_7" at 749,408 size 70x22; FormatPattern 9.9; Unit  
      ProcessValue <- "16_AQ_Data_R2_SPR_AQ_98"
   TextField "Text field_14" at 481,408 size 220x22; Text 'Spare'
   TextField "Text field_15" at 429,368 size 53x22; Text 'QW96'
   TextField "Text field_16" at 428,408 size 53x22; Text 'QW98'
   Group "Group" at 455,41 size 373x50
   Button "HmiScreenItemData_8" at 469,45 size 355x40; TextOn 'Back'; TextOff 'Text'
   TextField "Screen title" at 455,41 size 373x50; Text 'Screen title'

screen "GCU Analogue Outputs" 1280x800, template "Template"
   on GenerateScreen: "TitleUpdater"()
   Button "HmiScreenItemData_1" at 1,1 size 150x43; TextOn 'Back'; TextOff 'Commissioning'
      on Release: ActivateScreen("Commissioning Main Page", 0)
   Button "Button_15" at 34,732 size 100x35; TextOn 'BWTS Digital Inputs'; TextOff 'Back'
      on Click: ActivateScreen("BC Analogue Inputs", 0)
   AlarmView "Alarm view_1" at 0,777 size 1280x23
   TextField "Text field_90" at 750,328 size 64x20; Text 'Reading'
   TextField "Text field_41" at 553,328 size 89x20; Text 'Description'
   TextField "Text field_43" at 437,328 size 37x20; Text 'AO'
   TextField "Text field_52" at 437,295 size 336x26; Text 'GCU Control System PLC (Rack 3)'
   TextField "Text field_4" at 481,444 size 220x22; Text 'Spare'
   IOField "I/O field_4" at 749,446 size 70x22; FormatPattern 9999
      ProcessValue <- "16_AQ_Data_R3_SPR_AQ_804"
   TextField "Text field_8" at 428,444 size 53x22; Text 'QW804'
   TextField "Text field_9" at 481,368 size 220x22; Text 'CV405 GAS VENT POSITION'
   TextField "Text field_12" at 480,482 size 220x22; Text 'Spare'
   IOField "I/O field_5" at 749,481 size 70x22; FormatPattern 9999
      ProcessValue <- "16_AQ_Data_R3_SPR_AQ_806"
   TextField "Text field_13" at 427,482 size 53x22; Text 'QW806'
   Button "Button_7" at 716,442 size 29x26; TextOff '+'
      on Press: function_b14e0dd5("80_From_HMI_MAN_AQ_INC_804", 0)
      Visibility <- "82_To_HMI_CRNT_MODE_GCU"
   Button "Button_8" at 824,442 size 29x26; TextOff '-'
      on Press: function_b14e0dd5("80_From_HMI_MAN_AQ_DEC_804", 0)
      Visibility <- "82_To_HMI_CRNT_MODE_GCU"
   Button "Button_9" at 717,480 size 29x26; TextOff '+'
      on Press: function_b14e0dd5("80_From_HMI_MAN_AQ_INC_806", 0)
      Visibility <- "82_To_HMI_CRNT_MODE_GCU"
   Button "Button_10" at 825,480 size 29x26; TextOff '-'
      on Press: function_b14e0dd5("80_From_HMI_MAN_AQ_DEC_806", 0)
      Visibility <- "82_To_HMI_CRNT_MODE_GCU"
   Button "Button_11" at 716,364 size 29x26; TextOff '+'
      on Press: function_b14e0dd5("80_From_HMI_MAN_AQ_INC_800", 0)
      Visibility <- "82_To_HMI_CRNT_MODE_GCU"
   Button "Button_12" at 824,364 size 29x26; TextOff '-'
      on Press: function_b14e0dd5("80_From_HMI_MAN_AQ_DEC_800", 0)
      Visibility <- "82_To_HMI_CRNT_MODE_GCU"
   Button "Button_13" at 717,405 size 29x26; TextOff '+'
      on Press: function_b14e0dd5("80_From_HMI_MAN_AQ_INC_802", 0)
      Visibility <- "82_To_HMI_CRNT_MODE_GCU"
   Button "Button_14" at 825,405 size 29x26; TextOff '-'
      on Press: function_b14e0dd5("80_From_HMI_MAN_AQ_DEC_802", 0)
      Visibility <- "82_To_HMI_CRNT_MODE_GCU"
   IOField "I/O field_6" at 750,368 size 70x22; FormatPattern 999; Unit   %
      ProcessValue <- "16_AQ_Data_CV405_CNTRL"
   IOField "I/O field_7" at 751,408 size 70x22; FormatPattern 9999; Unit  
      ProcessValue <- "16_AQ_Data_R3_SPR_AQ_802"
   TextField "Text field_14" at 481,408 size 220x22; Text 'Spare'
   TextField "Text field_15" at 429,368 size 53x22; Text 'QW800'
   TextField "Text field_16" at 428,408 size 53x22; Text 'QW802'
   Group "Group" at 455,41 size 373x50
   Button "HmiScreenItemData_8" at 469,45 size 355x40; TextOn 'Back'; TextOff 'Text'
   TextField "Screen title" at 455,41 size 373x50; Text 'Screen title'

screen "BWT Analogue Outputs" 1280x800, template "Template"
   on GenerateScreen: "TitleUpdater"()
   Button "HmiScreenItemData_1" at 1,1 size 150x43; TextOn 'Back'; TextOff 'Commissioning'
      on Release: ActivateScreen("Commissioning Main Page", 0)
   TextField "Text field_90" at 799,171 size 64x20; Text 'Reading'
   TextField "Text field_41" at 602,171 size 89x20; Text 'Description'
   TextField "Text field_43" at 486,171 size 37x20; Text 'AO'
   TextField "Text field_52" at 486,138 size 340x26; Text 'BWT Control System PLC (Rack 3)'
   TextField "Text field_4" at 530,287 size 220x22; Text 'Main Fuel Reg Valve Control'
   IOField "I/O field_4" at 798,289 size 70x22; FormatPattern 9999; Unit %
      ProcessValue <- "16_AQ_Data_CV203_CNTRL"
   TextField "Text field_8" at 477,287 size 53x22; Text 'QW100'
   TextField "Text field_9" at 530,211 size 220x22; Text 'Spare'
   TextField "Text field_12" at 529,325 size 220x22; Text 'Main Atom Air Reg Valve Control'
   IOField "I/O field_5" at 798,324 size 70x22; FormatPattern 9999; Unit %
      ProcessValue <- "16_AQ_Data_CV111_CNTRL"
   TextField "Text field_13" at 476,325 size 53x22; Text 'QW102'
   Button "Button_7" at 765,285 size 29x26; TextOff '+'
      on Press: function_b14e0dd5("80_From_HMI_MAN_AQ_INC_100(1)", 0)
      Visibility <- "82_To_HMI_CRNT_MODE_IGG"
   Button "Button_8" at 873,285 size 29x26; TextOff '-'
      on Press: function_b14e0dd5("80_From_HMI_MAN_AQ_DEC_100(1)", 0)
      Visibility <- "82_To_HMI_CRNT_MODE_IGG"
   Button "Button_9" at 766,323 size 29x26; TextOff '+'
      on Press: function_b14e0dd5("80_From_HMI_MAN_AQ_INC_102", 0)
      Visibility <- "82_To_HMI_CRNT_MODE_IGG"
   Button "Button_10" at 874,323 size 29x26; TextOff '-'
      on Press: function_b14e0dd5("80_From_HMI_MAN_AQ_DEC_102", 0)
      Visibility <- "82_To_HMI_CRNT_MODE_IGG"
   Button "Button_11" at 765,207 size 29x26; TextOff '+'
      on Click: SetBit("80_From_HMI_MAN_AQ_INC_96")
      Visibility <- "82_To_HMI_CRNT_MODE_IGG"
   Button "Button_12" at 873,207 size 29x26; TextOff '-'
      on Click: SetBit("80_From_HMI_MAN_AQ_DEC_96")
      Visibility <- "82_To_HMI_CRNT_MODE_IGG"
   Button "Button_13" at 766,248 size 29x26; TextOff '+'
      on Click: SetBit("80_From_HMI_MAN_AQ_INC_98")
      Visibility <- "82_To_HMI_CRNT_MODE_IGG"
   Button "Button_14" at 874,248 size 29x26; TextOff '-'
      on Click: SetBit("80_From_HMI_MAN_AQ_DEC_98")
      Visibility <- "82_To_HMI_CRNT_MODE_IGG"
   IOField "I/O field_6" at 799,211 size 70x22; FormatPattern 9.9; Unit  
      ProcessValue <- "16_AQ_Data_R2_SPR_AQ_96"
   IOField "I/O field_7" at 800,251 size 70x22; FormatPattern 9.9; Unit  
      ProcessValue <- "16_AQ_Data_R2_SPR_AQ_98"
   TextField "Text field_14" at 530,251 size 220x22; Text 'Spare'
   TextField "Text field_15" at 478,211 size 53x22; Text 'QW96'
   TextField "Text field_16" at 477,251 size 53x22; Text 'QW98'
   Button "Button_15" at 34,732 size 100x35; TextOn 'BWTS Digital Inputs'; TextOff 'Back'
      on Click: ActivateScreen("BC Analogue Inputs", 0)
   AlarmView "Alarm view_1" at 0,777 size 1280x23
   TextField "Text field_1" at 23,309 size 1188x123; Text 'Re - Work Required Througout This page'
   Group "Group" at 455,41 size 373x50
   Button "HmiScreenItemData_8" at 469,45 size 355x40; TextOn 'Back'; TextOff 'Text'
   TextField "Screen title" at 455,41 size 373x50; Text 'Screen title'

screen "BC Target Setpoints" 1280x800, template "Template"
   on GenerateScreen: "TitleUpdater"()
   Button "HmiScreenItemData_1" at 1,1 size 150x43; TextOn 'Back'; TextOff 'Commissioning'
      on Release: ActivateScreen("Commissioning Main Page", 0)
   AlarmView "Alarm view_1" at 0,777 size 1280x23
   TextField "Text field_25" at 394,430 size 407x22; Text 'PIT-113: IGG Main Atom Air Pressure Target'
   TextField "Text field_29" at 814,210 size 68x20; Text 'Setpoint'
   TextField "Text field_33" at 393,468 size 408x22; Text 'PIT-205: IGG Main Fuel Pressure Target'
   IOField "I/O field_58" at 816,468 size 60x22; Authorization "Parameter Change"; FormatPattern 999.99
      ProcessValue <- "84_Setpoints_PIT205_Target(1)"
   TextField "Text field_35" at 394,552 size 406x22; Text 'E-600: O2 Cargo Blanketing Target'
   TextField "Text field_65" at 394,236 size 411x22; Text 'PIT-402: IG Outlet Pressure Pilot Target'
   TextField "Text field_67" at 394,274 size 410x22; Text 'PIT-402: IG Outlet Pressure Main Target'
   TextField "Text field_69" at 395,313 size 407x22; Text 'PIT-402: IG Outlet Pressure Post Target Start'
   TextField "Text field_71" at 395,352 size 406x22; Text 'PIT-402: IG Outlet Pressure Post Target Maximum'
   TextField "Text field_73" at 395,391 size 407x22; Text 'FD-001: Igniter Target'
   TextField "Text field_42" at 394,210 size 89x20; Text 'Description'
   IOField "I/O field_128" at 816,236 size 60x22; Authorization "Parameter Change"; FormatPattern 999.9
      ProcessValue <- "84_Setpoints_PIT402_Pilot_Target(1)"
   IOField "I/O field_133" at 816,274 size 60x22; Authorization "Parameter Change"; FormatPattern 999.9
      ProcessValue <- "84_Setpoints_PIT402_Main_Target(1)"
   IOField "I/O field_138" at 816,313 size 60x22; Authorization "Parameter Change"; FormatPattern 999.9
      ProcessValue <- "84_Setpoints_PIT402_Post_Target_Start"
   IOField "I/O field_53" at 816,430 size 60x22; Authorization "Parameter Change"; FormatPattern 999.9
      ProcessValue <- "84_Setpoints_PIT113_Pilot_Target(1)"
   IOField "I/O field_148" at 816,391 size 60x22; Authorization "Parameter Change"; FormatPattern 999.9
      ProcessValue <- "84_Setpoints_FD001_Min"
   IOField "I/O field_64" at 816,552 size 60x22; Authorization "Parameter Change"; FormatPattern 99.9
      ProcessValue <- "84_Setpoints_E600_CB_Target"
   TextField "Text field_53" at 393,184 size 213x26; Text 'IGG Target Setpoints'
   IOField "I/O field_5" at 815,352 size 60x22; Authorization "Parameter Change"; FormatPattern 999.9
      ProcessValue <- "84_Setpoints_PIT401_Post_Target_Max"
   TextField "Text field_1" at 394,510 size 406x22; Text 'E-600: O2 Ballast Water Treatment Target'
   IOField "I/O field_2" at 816,510 size 60x22; Authorization "Parameter Change"; FormatPattern 9.99
      ProcessValue <- "84_Setpoints_E600_BWT_Target"
   TextField "Text field_2" at 394,595 size 406x22; Text 'PIT-402 Target Ramp Time (s)'
   IOField "I/O field_1" at 816,595 size 60x22; Authorization "Parameter Change"; FormatPattern 99
      ProcessValue <- "19_AUTO_CMNDS_Data_PIT402_Target"
   Group "Group" at 455,41 size 373x50
   Button "HmiScreenItemData_8" at 469,45 size 355x40; TextOn 'Back'; TextOff 'Text'
   TextField "Screen title" at 455,41 size 373x50; Text 'Screen title'

